                 //check for max outlier
                 //calculate border for outlier
                 #statBorderOutlier := #statQuartil75 + #rangeOutlier * #statDeltaQuartil;
                 //search in array for values outside the border 
                 FOR #statCounter := UDINT_TO_INT(#statNumberOfElements - 1) TO 0 BY -1 DO
                   #statRetVal := MOVE_BLK_VARIANT(SRC := #array, COUNT := 1, SRC_INDEX := #statCounter, DEST_INDEX := 0, DEST => #tempValueInt);
                   IF #statRetVal <> 0
                   THEN
                     #status := INT_TO_WORD(#statRetVal);
                     #statusID := #ID_INTERNAL;
                     #statError := true;
                     GOTO EndOfBlock;
                   END_IF;
                   IF #tempValueInt > #statBorderOutlier
                   THEN
                     //detected a value as outlier, check next value
                     ;
                   ELSE
                     //all outlier detected. Calulate new Max Value in range and calulate outliers in %
                     #statOutlierMax := INT_TO_REAL((100 * (UDINT_TO_INT(#statNumberOfElements) - #statCounter - 1))) / UDINT_TO_REAL(#statNumberOfElements);
                     #statMaxNew := #tempValueInt;
                     EXIT;
                   END_IF;
                 END_FOR;
               END_IF;

               //done
               #statDone := TRUE;
             END_IF;
           END_REGION ;

         ELSIF TypeOfElements(#array) = UInt
         THEN

           REGION Type is UINT
             //Type is UInt 
             //Sort array
             #instLGF_ShellSortUInt(error => #statError,
                                    statusID => #tempStatusID,
                                    status => #tempStatus,
                                    variantArray := #array);

             IF #statError = true
             THEN
               IF #tempStatusID > 1
               THEN
                 #statusID := #ID_INTERNAL;
               ELSE
                 #statusID := #ID_SORT;
                 #status := #tempStatus;
               END_IF;
               GOTO EndOfBlock;
             END_IF;

             //Identify max and min value
             #statRetVal := MOVE_BLK_VARIANT(SRC := #array, COUNT := 1, SRC_INDEX := 0, DEST_INDEX := 0, DEST => #tempMinUint);
             IF #statRetVal <> 0
             THEN
               #status := INT_TO_WORD(#statRetVal);
               #statusID := #ID_INTERNAL;
               #statError := true;
               GOTO EndOfBlock;
             END_IF;
             #statRetVal := MOVE_BLK_VARIANT(SRC := #array, COUNT := 1, SRC_INDEX := UDINT_TO_INT(#statNumberOfElements - 1), DEST_INDEX := 0, DEST => #tempMaxUint);
             IF #statRetVal <> 0
             THEN
               #status := INT_TO_WORD(#statRetVal);
               #statusID := #ID_INTERNAL;
               #statError := true;
               GOTO EndOfBlock;
             END_IF;
             #statMax := #tempMaxUint;
             #statMin := #tempMinUint;

             //calculate median (Q50)
             IF #statEven = true
             THEN
               // if n is even -> calculate MEDIAN = (x(n/2)+x(n/2+1))/2
               #statRetVal := MOVE_BLK_VARIANT(SRC := #array, COUNT := 1, SRC_INDEX := UDINT_TO_INT(#statNumberOfElements / 2), DEST_INDEX := 0, DEST => #tempValueUint);
               IF #statRetVal <> 0
               THEN
                 #status := INT_TO_WORD(#statRetVal);
                 #statusID := #ID_INTERNAL;
                 #statError := true;
                 GOTO EndOfBlock;
               END_IF;
               #statRetVal := MOVE_BLK_VARIANT(SRC := #array, COUNT := 1, SRC_INDEX := UDINT_TO_INT(#statNumberOfElements / 2) - 1, DEST_INDEX := 0, DEST => #tempValueUint1);
               IF #statRetVal <> 0
               THEN
                 #status := INT_TO_WORD(#statRetVal);
                 #statusID := #ID_INTERNAL;
                 #statError := true;
                 GOTO EndOfBlock;
               END_IF;
               #statMedian := (#tempValueUint + #tempValueUint1) / 2;
             ELSE
               // if n is odd -> MEDIAN = x(n+1/2)
               #statRetVal := MOVE_BLK_VARIANT(SRC := #array, COUNT := 1, SRC_INDEX := UDINT_TO_INT(#statNumberOfElements / 2), DEST_INDEX := 0, DEST => #tempValueUint);
               IF #statRetVal <> 0
               THEN
                 #status := INT_TO_WORD(#statRetVal);
                 #statusID := #ID_INTERNAL;
                 #statError := true;
                 GOTO EndOfBlock;
               END_IF;
               #statMedian := #tempValueUint;
             END_IF;

             //calculate 1.quartil (Q25)
             // q1 = x(k) with  k=(n+3)/4 
             #statK := (((UDINT_TO_REAL(#statNumberOfElements + 3)) / 4.0)) - 1;
             #statRetVal := MOVE_BLK_VARIANT(SRC := #array, COUNT := 1, SRC_INDEX := TRUNC(#statK), DEST_INDEX := 0, DEST => #tempValueUint);
             IF #statRetVal <> 0
             THEN
               #status := INT_TO_WORD(#statRetVal);
               #statError := true;
               GOTO EndOfBlock;
             END_IF;
             #statRetVal := MOVE_BLK_VARIANT(SRC := #array, COUNT := 1, SRC_INDEX := TRUNC(#statK) + 1, DEST_INDEX := 0, DEST => #tempValueUint1);
             IF #statRetVal <> 0
             THEN
               #status := INT_TO_WORD(#statRetVal);
               #statusID := #ID_INTERNAL;
               #statError := true;
               GOTO EndOfBlock;
             END_IF;

             #statQuartil25 := #tempValueUint + FRAC_REAL(#statK) * (#tempValueUint1 - #tempValueUint);
             //calculate 3.quartil (Q75)
             //q3 = x(n+1-k) with k=(3n+1)/4
             #statK := ((3 * UDINT_TO_REAL(#statNumberOfElements) + 1) / 4) - 1;
             #statRetVal := MOVE_BLK_VARIANT(SRC := #array, COUNT := 1, SRC_INDEX := TRUNC(#statK), DEST_INDEX := 0, DEST => #tempValueUint);
             IF #statRetVal <> 0
             THEN
               #status := INT_TO_WORD(#statRetVal);
               #statusID := #ID_INTERNAL;
               #statError := true;
               GOTO EndOfBlock;
             END_IF;
             #statRetVal := MOVE_BLK_VARIANT(SRC := #array, COUNT := 1, SRC_INDEX := TRUNC(#statK) + 1, DEST_INDEX := 0, DEST => #tempValueUint1);
             IF #statRetVal <> 0
             THEN
               #status := INT_TO_WORD(#statRetVal);
               #statusID := #ID_INTERNAL;
               #statError := true;
               GOTO EndOfBlock;
             END_IF;

             #statQuartil75 := #tempValueUint + FRAC_REAL(#statK) * (#tempValueUint1 - #tempValueUint);

             //only if RANGE_OUTLIER <> 0
             IF #rangeOutlier <> 0
             THEN

               //calculate Delta Q75-Q25
               #statDeltaQuartil := #statQuartil75 - #statQuartil25;

               //calculate border for outlier
               #statBorderOutlier := #statQuartil25 - #rangeOutlier * #statDeltaQuartil;
               //search in array for values outside the border
               FOR #statCounter := 0 TO UDINT_TO_INT(#statNumberOfElements - 1) DO
                 #statRetVal := MOVE_BLK_VARIANT(SRC := #array, COUNT := 1, SRC_INDEX := #statCounter, DEST_INDEX := 0, DEST => #tempValueUint);
                 IF #statRetVal <> 0
                 THEN
                   #status := INT_TO_WORD(#statRetVal);
                   #statusID := #ID_INTERNAL;
                   #statError := true;
                   GOTO EndOfBlock;
                 END_IF;
                 IF #tempValueUint < #statBorderOutlier
                 THEN
                   //detected a value as outlier, check next value
                   ;
                 ELSE
                   //all outlier detected. Calulate new Min Value in range and calulate outliers in %
                   #statOutlierMin := INT_TO_REAL((100 * #statCounter)) / UDINT_TO_REAL(#statNumberOfElements);
                   #statMinNew := #tempValueUint;
                   EXIT;
                 END_IF;

               END_FOR;

               //check for max outlier
               #statBorderOutlier := #statQuartil75 + #rangeOutlier * #statDeltaQuartil;

               FOR #statCounter := UDINT_TO_INT(#statNumberOfElements - 1) TO 0 BY -1 DO
                 #statRetVal := MOVE_BLK_VARIANT(SRC := #array, COUNT := 1, SRC_INDEX := #statCounter, DEST_INDEX := 0, DEST => #tempValueUint);
                 IF #statRetVal <> 0
                 THEN
                   #status := INT_TO_WORD(#statRetVal);
                   #statusID := #ID_INTERNAL;
                   #statError := true;
                   GOTO EndOfBlock;
                 END_IF;
                 IF #tempValueUint > #statBorderOutlier
                 THEN
                   //detected a value as outlier, check next value
                   ;
                 ELSE
                   //all outlier detected. Calulate new Max Value in range and calulate outliers in %
                   #statOutlierMax := INT_TO_REAL((100 * (UDINT_TO_INT(#statNumberOfElements) - #statCounter - 1))) / UDINT_TO_REAL(#statNumberOfElements);
                   #statMaxNew := #tempValueUint;
                   EXIT;
                 END_IF;
               END_FOR;
             END_IF;
             //done
             #statDone := TRUE;

           END_REGION ;

         ELSIF TypeOfElements(#array) = Real
         THEN

           REGION Type of Array is REAL

             //Type is Real
             //Sort array
             #instLGF_ShellSortReal(error => #statError,
                                    statusID => #tempStatusID,
                                    status => #tempStatus,
                                    variantArray := #array);

             IF #statError = true
             THEN
               IF #tempStatusID > 1
               THEN
                 #statusID := #ID_INTERNAL;
               ELSE
                 #statusID := #ID_SORT;
                 #status := #tempStatus;
               END_IF;
               GOTO EndOfBlock;
             END_IF;

             //Identify max and min value
             #statRetVal := MOVE_BLK_VARIANT(SRC := #array, COUNT := 1, SRC_INDEX := 0, DEST_INDEX := 0, DEST => #statMin);
             IF #statRetVal <> 0
             THEN
               #status := INT_TO_WORD(#statRetVal);
               #statusID := #ID_INTERNAL;
               #statError := true;
               GOTO EndOfBlock;
             END_IF;
             #statRetVal := MOVE_BLK_VARIANT(SRC := #array, COUNT := 1, SRC_INDEX := UDINT_TO_INT(#statNumberOfElements - 1), DEST_INDEX := 0, DEST => #statMax);
             IF #statRetVal <> 0
             THEN
               #status := INT_TO_WORD(#statRetVal);
               #statusID := #ID_INTERNAL;
               #statError := true;
               GOTO EndOfBlock;
             END_IF;

             //calculate median (Q50)
             IF #statEven = true
             THEN
               // if n is even -> calculate MEDIAN = (x(n/2)+x(n/2+1))/2
               #statRetVal := MOVE_BLK_VARIANT(SRC := #array, COUNT := 1, SRC_INDEX := UDINT_TO_INT(#statNumberOfElements / 2), DEST_INDEX := 0, DEST => #tempValueReal);
               IF #statRetVal <> 0
               THEN
                 #status := INT_TO_WORD(#statRetVal);
                 #statusID := #ID_INTERNAL;
                 #statError := true;
                 GOTO EndOfBlock;
               END_IF;
               #statRetVal := MOVE_BLK_VARIANT(SRC := #array, COUNT := 1, SRC_INDEX := UDINT_TO_INT(#statNumberOfElements / 2) - 1, DEST_INDEX := 0, DEST => #tempValueReal1);
               IF #statRetVal <> 0
               THEN
                 #status := INT_TO_WORD(#statRetVal);
                 #statusID := #ID_INTERNAL;
                 #statError := true;
                 GOTO EndOfBlock;
               END_IF;
               #statMedian := (#tempValueReal + #tempValueReal1) / 2;
             ELSE
               // if n is odd -> MEDIAN = x(n+1/2)
               #statRetVal := MOVE_BLK_VARIANT(SRC := #array, COUNT := 1, SRC_INDEX := UDINT_TO_INT(#statNumberOfElements / 2), DEST_INDEX := 0, DEST => #tempValueReal);
               IF #statRetVal <> 0
               THEN
                 #status := INT_TO_WORD(#statRetVal);
                 #statusID := #ID_INTERNAL;
                 #statError := true;
                 GOTO EndOfBlock;
               END_IF;
               #statMedian := #tempValueReal;
             END_IF;

             //calculate 1.quartil (Q25)
             // q1 = x(k) with  k=(n+3)/4 
             #statK := (((UDINT_TO_REAL(#statNumberOfElements + 3)) / 4.0)) - 1;
             #statRetVal := MOVE_BLK_VARIANT(SRC := #array, COUNT := 1, SRC_INDEX := TRUNC(#statK), DEST_INDEX := 0, DEST => #tempValueReal);
             IF #statRetVal <> 0
             THEN
               #status := INT_TO_WORD(#statRetVal);
               #statusID := #ID_INTERNAL;
               #statError := true;
               GOTO EndOfBlock;
             END_IF;
             #statRetVal := MOVE_BLK_VARIANT(SRC := #array, COUNT := 1, SRC_INDEX := TRUNC(#statK) + 1, DEST_INDEX := 0, DEST => #tempValueReal1);
             IF #statRetVal <> 0
             THEN
               #status := INT_TO_WORD(#statRetVal);
               #statusID := #ID_INTERNAL;
               #statError := true;
               GOTO EndOfBlock;
             END_IF;
             #statQuartil25 := #tempValueReal + FRAC_REAL(#statK) * (#tempValueReal1 - #tempValueReal);

             //calculate 3.quartil (Q75)
             //q3 = x(n+1-k) with k=(3n+1)/4
             #statK := ((3 * UDINT_TO_REAL(#statNumberOfElements) + 1) / 4) - 1;
             #statRetVal := MOVE_BLK_VARIANT(SRC := #array, COUNT := 1, SRC_INDEX := TRUNC(#statK), DEST_INDEX := 0, DEST => #tempValueReal);
             IF #statRetVal <> 0
             THEN
               #status := INT_TO_WORD(#statRetVal);
               #statusID := #ID_INTERNAL;
               #statError := true;
               GOTO EndOfBlock;
             END_IF;
             #statRetVal := MOVE_BLK_VARIANT(SRC := #array, COUNT := 1, SRC_INDEX := TRUNC(#statK) + 1, DEST_INDEX := 0, DEST => #tempValueReal1);
             IF #statRetVal <> 0
             THEN
               #status := INT_TO_WORD(#statRetVal);
               #statusID := #ID_INTERNAL;
               #statError := true;
               GOTO EndOfBlock;
             END_IF;
             #statQuartil75 := #tempValueReal + FRAC_REAL(#statK) * (#tempValueReal1 - #tempValueReal);

             //only if RANGE_OUTLIER <> 0
             IF #rangeOutlier <> 0
             THEN

               //calculate Delta Q75-Q25
               #statDeltaQuartil := #statQuartil75 - #statQuartil25;

               //calculate border for outlier
               #statBorderOutlier := #statQuartil25 - #rangeOutlier * #statDeltaQuartil;
               FOR #statCounter := 0 TO UDINT_TO_INT(#statNumberOfElements - 1) DO
                 #statRetVal := MOVE_BLK_VARIANT(SRC := #array, COUNT := 1, SRC_INDEX := #statCounter, DEST_INDEX := 0, DEST => #tempValueReal);
                 IF #statRetVal <> 0
                 THEN
                   #status := INT_TO_WORD(#statRetVal);
                   #statusID := #ID_INTERNAL;
                   #statError := true;
                   GOTO EndOfBlock;
                 END_IF;
                 IF #tempValueReal < #statBorderOutlier
                 THEN
                   //detected a value as outlier, check next value
                   ;
                 ELSE
                   //all outlier detected. Calulate new Min Value in range and calulate outliers in %
                   #statOutlierMin := INT_TO_REAL((100 * #statCounter)) / UDINT_TO_REAL(#statNumberOfElements);
                   #statMinNew := #tempValueReal;
                   EXIT;
                 END_IF;

               END_FOR;

               //check for max outlier
               //calculate border for outlier
               #statBorderOutlier := #statQuartil75 + #rangeOutlier * #statDeltaQuartil;
               FOR #statCounter := UDINT_TO_INT(#statNumberOfElements - 1) TO 0 BY -1 DO
                 #statRetVal := MOVE_BLK_VARIANT(SRC := #array, COUNT := 1, SRC_INDEX := #statCounter, DEST_INDEX := 0, DEST => #tempValueReal);
                 IF #statRetVal <> 0
                 THEN
                   #status := INT_TO_WORD(#statRetVal);
                   #statusID := #ID_INTERNAL;
                   #statError := true;
                   GOTO EndOfBlock;
                 END_IF;
                 IF #tempValueReal > #statBorderOutlier
                 THEN
                   //detected a value as outlier, check next value
                   ;
                 ELSE
                   //all outlier detected. Calulate new Max Value in range and calulate outliers in %
                   #statOutlierMax := INT_TO_REAL((100 * (UDINT_TO_INT(#statNumberOfElements) - #statCounter - 1))) / UDINT_TO_REAL(#statNumberOfElements);
                   #statMaxNew := #tempValueReal;
                   EXIT;
                 END_IF;
               END_FOR;
             END_IF;
             //done
             #statDone := TRUE;

           END_REGION ;

         ELSE
           #statError := true;
           #status := #STATUS_WRONG_DATATYPE;
         END_IF;
         //calculate Skewness
         //S= ((Q25 + Q75)-2*Q50) / (Q75 - Q25)
         #skewness := (#statQuartil75 + #statQuartil25 - 2.0 * #statMedian) / (#statQuartil75 - #statQuartil25);

         //write output values
         IF #rangeOutlier <> 0
         THEN
           #min := #statMinNew;
           #max := #statMaxNew;
         ELSE
           #min := #statMin;
           #max := #statMax;
         END_IF;

         #q25 := #statQuartil25;
         #median := #statMedian;
         #q75 := #statQuartil75;
         #outlierMin := #statOutlierMin;
         #outlierMax := #statOutlierMax;
         GOTO EndOfBlock;

       END_IF;
     ELSE
       #statError := true;
       #status := #STATUS_NO_ARRAY;
     END_IF;


   END_REGION

   REGION Write Outputs
     //Error occured in request


   EndOfBlock:
     IF #statError
     THEN
       #statDone := FALSE;
       #statBusy := FALSE;
       //Request finished
     ELSIF #statDone
     THEN
       #statBusy := FALSE;
       #statError := FALSE;
       #status := #STATUS_EXECUTION_FINISHED;

       //Request in execution
     ELSE
       #status := #STATUS_SUBSEQUENT_CALL;
     END_IF;


     //Write static values (done,busy,error) to outputs
     #done := #statDone;
     #busy := #statBusy;
     #error := #statError;
     //----------------------------------------------------------------------------------------------

   END_REGION ;
END_FUNCTION_BLOCK

FUNCTION_BLOCK "LGF_Histogram"   // FB10011, SCL
{ S7_Optimized_Access := 'TRUE' }
VERSION : 0.1
   VAR_INPUT
      execute : Bool;   // Rising edge starts action once
      NumberOfClasses : UInt;   // Number of desired classes.
   END_VAR
   VAR_OUTPUT
      busy : Bool;   // TRUE: FB is not finished and new output values can be expected
      done : Bool;   // TRUE: Commanded action has been completed successfully
      error : Bool;   // Rising edge informs that an error occurred during the execution of
      status : Word := 16#7000;   // Current status of FB
      statusID : UInt := 1;   // Current statusID of FB
      histValues : Array[0..1, 0..14] of Real;   // Outputs the calculated values in a two-dimensional array
      axis : Array[0..3] of Real;   // Specifies the axis values
      classWidth : Real;   // Returns the calculated class width.
   END_VAR
   VAR_IN_OUT
      "array" : Variant;
   END_VAR
   VAR
      statBusy : Bool;   // Static value for output busy
      statDone : Bool;   // Static value for output done
      statError : Bool;   // Static value for output error
      statExecuteOld : Bool;   // Old value of execute for edge detection
      instLGF_ShellSortInt : "LGF_ShellSortInt";   // Instance of LG_ShellSortInt
      instLGF_ShellSortReal : "LGF_ShellSortReal";   // Instance of LG_ShellSortReal
      instLGF_ShellSortUInt : "LGF_ShellSortUInt";   // Instance of LG_ShellSortUInt
      statMin : Real;   // Static value for min
      statMax : Real;   // Static value for max
      statNumberOfElements : UDInt;   // Static value for number of elements
      statType : Int;   // Static value for type
      statAverage : Real;   // Static value for average
      statDeviation : Real;   // Static value for deviation
      statCounter : Int;   // Static value for counter
      statWidth : Real;   // Static value for width
      statFrequencyValues : Int;   // Static value for frequency values
      statI : Int;   // Static value for I
      statIold : Int := 0;   // Static value for I old
      statBound : Real;   // Static value for bound
      statMaxFrequency : Int;   // Static value for max frequency
      statHistFrequencyAbs : Array[0..14] of Int;   // Static array for history frequency absolute
      statHistFrequencyRel : Array[0..14] of Real;   // Static array for history frequency relative
      statHistMiddleOfClass : Array[0..14] of Real;   // Static array for history middle of class
   END_VAR
   VAR_TEMP
      tempError : Bool;   // Temporary error
      tempStatusID : UInt;   // Temporary status ID
      tempStatus : Word;   // Temporary status
      tempRetVal : Int;   // Temporary RetVal
      tempValueInt : Int;   // Temporary value for calculation
      tempValueUint : UInt;   // Temporary value for calculation
      tempValueReal : Real;   // Temporary value for calculation
      tempMinInt : Int;   // Temporary value for min INT
      tempMaxInt : Int;   // Temporary value for max INT
      tempMinUint : UInt;   // Temporary value for min UINT
      tempMaxUint : UInt;   // Temporary value for max UINT
   END_VAR
   VAR CONSTANT
      STATUS_EXECUTION_FINISHED : Word := 16#0000;   // Status: Execution finished without errors
      STATUS_NO_CALL : Word := 16#7000;   // Status: No call of FB
      STATUS_FIRST_CALL : Word := 16#7001;   // Status: First call of FB after enabling
      STATUS_SUBSEQUENT_CALL : Word := 16#7002;   // Status: Subsequent call of FB
      STATUS_WRONG_DATATYPE : Word := 16#9100;   // Status: Wrong data type
      STATUS_WRONG_NO_CLASSES : Word := 16#9101;   // Status: Wrong number of classes
      STATUS_NO_ARRAY : Word := 16#9102;   // Status: No array
      TYPE_INT : Int := 0;   // TYPE: INT
      TYPE_UINT : Int := 1;   // TYPE: UINT
      TYPE_REAL : Int := 2;   // TYPE: REAL
      ID_INTERNAL : UInt := 1;   // Status ID: Internal error
      ID_MOVE_BLK : UInt := 2;   // Status ID: Function MOVE_BLK
      ID_SORT : UInt := 3;   // Status ID: Error sorting
   END_VAR
BEGIN
   //=============================================================================
   // SIEMENS AG
   // (c)Copyright 2017
   //-----------------------------------------------------------------------------
   // Library:       LGF (Library General Functions)
   // Tested with:   CPU1212C DC/DC/DC FW:V4.2
   // Engineering:   TIA Portal V15.1 
   // Restrictions:  -
   // Requirements:  PLC (S7-1200 / S7-1500)
   // Functionality: calculate from measurement list all values for creating
   //                a histogramm with WinCC
   //-----------------------------------------------------------------------------
   // Change log table:
   // Version  Date        In charge / Changes applied
   // 01.00.00 23.11.2018  Siemens Industry Online Support
   //                      First released version
   //=============================================================================

   //Check if FB is triggered
   //Too many classes on input. MAX = 15 Classes

   //FB is active
   IF #execute
     AND NOT #statExecuteOld
     AND NOT #statBusy
   THEN
     //Functionality is busy
     #statBusy := TRUE;

     //Reset other outputs
     #statError := FALSE;
     #status := #STATUS_FIRST_CALL;

     //Reset statics
     FILL_BLK(IN := 0,
              COUNT := 15,
              OUT => #statHistFrequencyAbs[0]);
     FILL_BLK(IN := 0,
              COUNT := 15,
              OUT => #statHistFrequencyRel[0]);
     FILL_BLK(IN := 0,
              COUNT := 15,
              OUT => #statHistMiddleOfClass[0]);
     #statI := 0;
     #statFrequencyValues := 0;
     #statIold := 0;

     #statExecuteOld := #execute;
     #statMaxFrequency := 0;

     GOTO EndOfBlock;
     //FB is currently inactive
   ELSIF NOT #execute
     AND NOT #statBusy
   THEN
     //Error outputs are reset with falling edge of enable input
     #statError := FALSE;

     //Done and busy are reset with falling edge of enable input
     #statDone := FALSE;
     #statBusy := FALSE;

     //Write outputs
     #status := #STATUS_NO_CALL;
     #statExecuteOld := #execute;

     GOTO EndOfBlock;
     //FB is currently executed and not finished
   ELSIF #statBusy
   THEN
     #statExecuteOld := #execute;

     //FB finished job
   ELSE
     #statExecuteOld := #execute;
     //Wait for start of functionality 
   END_IF;

   IF #statBusy = true
     AND #statError = false
   THEN

     REGION check Datatype of Array, sort and count the elements

       //count array elements
       #statNumberOfElements := CountOfElements(#array);

       //check number of classes
       IF (#NumberOfClasses > 15)
         OR (#NumberOfClasses < 1)
       THEN
         #statError := true;
         #status := #STATUS_WRONG_NO_CLASSES;
         #statusID := #ID_INTERNAL;
         GOTO EndOfBlock;
       END_IF;

       IF IS_ARRAY(#array)
       THEN
         //check which datatype is used
         IF TypeOfElements(#array) = Int
         THEN
           //Type is Int
           REGION Type of Array is INT
             //Sort array
             #instLGF_ShellSortInt(error => #statError,
                                   statusID => #tempStatusID,
                                   status => #tempStatus,
                                   variantArray := #array);
             IF #statError = true
             THEN
               IF #tempStatusID > 1
               THEN
                 #statusID := #ID_INTERNAL;
               ELSE
                 #statusID := #ID_SORT;
               END_IF;
               #status := #tempStatus;
               GOTO EndOfBlock;
             ELSE
               //Identify max and min value
               #tempRetVal := MOVE_BLK_VARIANT(SRC := #array, COUNT := 1, SRC_INDEX := 0, DEST_INDEX := 0, DEST => #tempMinInt);
               IF #tempRetVal <> 0
               THEN
                 #status := INT_TO_WORD(#tempRetVal);
                 #statusID := #ID_MOVE_BLK;
                 #statError := true;
                 GOTO EndOfBlock;
               END_IF;
               #tempRetVal := MOVE_BLK_VARIANT(SRC := #array, COUNT := 1, SRC_INDEX := UDINT_TO_INT(#statNumberOfElements - 1), DEST_INDEX := 0, DEST => #tempMaxInt);
               IF #tempRetVal <> 0
               THEN
                 #status := INT_TO_WORD(#tempRetVal);
                 #statusID := #ID_MOVE_BLK;
                 #statError := true;
                 GOTO EndOfBlock;
               END_IF;

               #statMin := INT_TO_REAL(#tempMinInt);
               #statMax := INT_TO_REAL(#tempMaxInt);

               //calculate classwidth
               #statWidth := (#statMax - #statMin) / #NumberOfClasses;
               #statBound := (#statMin + #statWidth);

               //search for all values
               FOR #statCounter := 0 TO UINT_TO_INT(#NumberOfClasses) - 1 DO

                 //Count Values for Class 
                 #tempRetVal := MOVE_BLK_VARIANT(SRC := #array, COUNT := 1, SRC_INDEX := 0, DEST_INDEX := 0, DEST => #tempValueInt);
                 IF #tempRetVal <> 0
                 THEN
                   #status := INT_TO_WORD(#tempRetVal);
                   #statusID := #ID_MOVE_BLK;
                   #statError := true;
                   GOTO EndOfBlock;
                 END_IF;
                 WHILE (#tempValueInt < #statBound)
                   AND #statI < #statNumberOfElements - 1 DO

                   IF #statI = #statNumberOfElements
                   THEN
                     EXIT;
                   END_IF;
                   #statI := #statI + 1;
                   #tempRetVal := MOVE_BLK_VARIANT(SRC := #array, COUNT := 1, SRC_INDEX := #statI, DEST_INDEX := 0, DEST => #tempValueInt);
                   IF #tempRetVal <> 0
                   THEN
                     #status := INT_TO_WORD(#tempRetVal);
                     #statusID := #ID_MOVE_BLK;
                     #statError := true;
                     GOTO EndOfBlock;
                   END_IF;
                 END_WHILE;

                 //the last value is not counted, because of rounding errors
                 IF #statI = #statNumberOfElements - 1
                 THEN
                   #statI := #statI + 1;
                 END_IF;

                 #statFrequencyValues := #statI - #statIold;
                 #statHistFrequencyAbs[#statCounter] := #statFrequencyValues;

                 #statHistFrequencyRel[#statCounter] := INT_TO_REAL(#statFrequencyValues) / UDINT_TO_REAL(#statNumberOfElements) * 100;

                 //Max values in one class for y-axis 
                 IF #statMaxFrequency < #statFrequencyValues
                 THEN
                   #statMaxFrequency := #statFrequencyValues;
                 END_IF;

                 #statBound := #statBound + #statWidth;
                 #statIold := #statI;
               END_FOR;
             END_IF;
           END_REGION

         ELSIF TypeOfElements(#array) = UInt
         THEN
           //Type is UInt 
           REGION Type of Array is UINT
             //Sort array
             #instLGF_ShellSortUInt(error => #statError,
                                    statusID => #tempStatusID,
                                    status => #tempStatus,
                                    variantArray := #array);
             IF #statError = true
             THEN
               IF #tempStatusID > 1
               THEN
                 #statusID := #ID_INTERNAL;
               ELSE
                 #statusID := #ID_SORT;
               END_IF;
               #status := #tempStatus;
               GOTO EndOfBlock;
             ELSE
               //Identify max and min value
               #tempRetVal := MOVE_BLK_VARIANT(SRC := #array, COUNT := 1, SRC_INDEX := 0, DEST_INDEX := 0, DEST => #tempMinUint);
               IF #tempRetVal <> 0
               THEN
                 #status := INT_TO_WORD(#tempRetVal);
                 #statusID := #ID_MOVE_BLK;
                 #statError := true;
                 GOTO EndOfBlock;
               END_IF;
               #tempRetVal := MOVE_BLK_VARIANT(SRC := #array, COUNT := 1, SRC_INDEX := UDINT_TO_INT(#statNumberOfElements - 1), DEST_INDEX := 0, DEST => #tempMaxUint);
               IF #tempRetVal <> 0
               THEN
                 #status := INT_TO_WORD(#tempRetVal);
                 #statusID := #ID_MOVE_BLK;
                 #statError := true;
                 GOTO EndOfBlock;
               END_IF;

               #statMin := UINT_TO_REAL(#tempMinUint);
               #statMax := UINT_TO_REAL(#tempMaxUint);

               //calculate classwidth
               #statWidth := (#statMax - #statMin) / #NumberOfClasses;
               #statBound := (#statMin + #statWidth);

               //search for all values
               FOR #statCounter := 0 TO UINT_TO_INT(#NumberOfClasses) - 1 DO

                 //Count Values for Class 
                 #tempRetVal := MOVE_BLK_VARIANT(SRC := #array, COUNT := 1, SRC_INDEX := 0, DEST_INDEX := 0, DEST => #tempValueUint);
                 IF #tempRetVal <> 0
                 THEN
                   #status := INT_TO_WORD(#tempRetVal);
                   #statusID := #ID_MOVE_BLK;
                   #statError := true;
                   GOTO EndOfBlock;

                 END_IF;
                 WHILE (#tempValueUint < #statBound)
                   AND #statI < #statNumberOfElements - 1 DO

                   IF #statI = #statNumberOfElements
                   THEN
                     EXIT;
                   END_IF;
                   #statI := #statI + 1;
                   #tempRetVal := MOVE_BLK_VARIANT(SRC := #array, COUNT := 1, SRC_INDEX := #statI, DEST_INDEX := 0, DEST => #tempValueUint);
                   IF #tempRetVal <> 0
                   THEN
                     #status := INT_TO_WORD(#tempRetVal);
                     #statusID := #ID_MOVE_BLK;
                     #statError := true;
                     GOTO EndOfBlock;
                   END_IF;
                 END_WHILE;

                 //the last value is not counted, because of rounding errors
                 IF #statI = #statNumberOfElements - 1
                 THEN
                   #statI := #statI + 1;
                 END_IF;

                 #statFrequencyValues := #statI - #statIold;
                 #statHistFrequencyAbs[#statCounter] := #statFrequencyValues;

                 #statHistFrequencyRel[#statCounter] := INT_TO_REAL(#statFrequencyValues) / UDINT_TO_REAL(#statNumberOfElements) * 100;

                 //Max values in one class for y-axis 
                 IF #statMaxFrequency < #statFrequencyValues
                 THEN
                   #statMaxFrequency := #statFrequencyValues;
                 END_IF;

                 #statBound := #statBound + #statWidth;
                 #statIold := #statI;
               END_FOR;

             END_IF;
           END_REGION

         ELSIF TypeOfElements(#array) = Real
         THEN
           //Type is Real
           REGION Type of Array is REAL
             //Sort array
             #instLGF_ShellSortReal(error => #statError,
                                    statusID => #tempStatusID,
                                    status => #tempStatus,
                                    variantArray := #array);
             IF #statError = true
             THEN
               IF #tempStatusID > 1
               THEN
                 #statusID := #ID_INTERNAL;
               ELSE
                 #statusID := #ID_SORT;
               END_IF;
               #status := #tempStatus;
               GOTO EndOfBlock;
             ELSE
               //Identify max and min value
               #tempRetVal := MOVE_BLK_VARIANT(SRC := #array, COUNT := 1, SRC_INDEX := 0, DEST_INDEX := 0, DEST => #statMin);
               IF #tempRetVal <> 0
               THEN
                 #status := INT_TO_WORD(#tempRetVal);
                 #statusID := #ID_MOVE_BLK;
                 #statError := true;
                 GOTO EndOfBlock;
               END_IF;
               #tempRetVal := MOVE_BLK_VARIANT(SRC := #array, COUNT := 1, SRC_INDEX := UDINT_TO_INT(#statNumberOfElements - 1), DEST_INDEX := 0, DEST => #statMax);
               IF #tempRetVal <> 0
               THEN
                 #status := INT_TO_WORD(#tempRetVal);
                 #statusID := #ID_MOVE_BLK;
                 #statError := true;
                 GOTO EndOfBlock;
               END_IF;
               //calculate classwidth
               #statWidth := (#statMax - #statMin) / #NumberOfClasses;
               #statBound := (#statMin + #statWidth);

               //search for all values
               FOR #statCounter := 0 TO UINT_TO_INT(#NumberOfClasses) - 1 DO

                 //Count Values for Class 
                 #tempRetVal := MOVE_BLK_VARIANT(SRC := #array, COUNT := 1, SRC_INDEX := 0, DEST_INDEX := 0, DEST => #tempValueReal);
                 IF #tempRetVal <> 0
                 THEN
                   #status := INT_TO_WORD(#tempRetVal);
                   #statusID := #ID_MOVE_BLK;
                   #statError := true;
                   GOTO EndOfBlock;
                 END_IF;
                 WHILE (#tempValueReal < #statBound)
                   AND #statI < #statNumberOfElements - 1 DO

                   IF #statI = #statNumberOfElements
                   THEN
                     EXIT;
                   END_IF;
                   #statI := #statI + 1;
                   #tempRetVal := MOVE_BLK_VARIANT(SRC := #array, COUNT := 1, SRC_INDEX := #statI, DEST_INDEX := 0, DEST => #tempValueReal);
                   IF #tempRetVal <> 0
                   THEN
                     #status := INT_TO_WORD(#tempRetVal);
                     #statusID := #ID_MOVE_BLK;
                     #statError := true;
                     GOTO EndOfBlock;
                   END_IF;
                 END_WHILE;

                 //the last value is not counted, because of rounding errors
                 IF #statI = #statNumberOfElements - 1
                 THEN
                   #statI := #statI + 1;
                 END_IF;

                 #statFrequencyValues := #statI - #statIold;
                 #statHistFrequencyAbs[#statCounter] := #statFrequencyValues;
                 #statHistFrequencyRel[#statCounter] := INT_TO_REAL(#statFrequencyValues) / UDINT_TO_REAL(#statNumberOfElements) * 100;

                 //Max values in one class for y-axis 
                 IF #statMaxFrequency < #statFrequencyValues
                 THEN
                   #statMaxFrequency := #statFrequencyValues;
                 END_IF;

                 #statBound := #statBound + #statWidth;
                 #statIold := #statI;
               END_FOR;
             END_IF;
             #statDone := true;
           END_REGION

         ELSE
           #statError := true;
           #status := #STATUS_WRONG_DATATYPE;
           GOTO EndOfBlock;
         END_IF;
       ELSE
         #statError := true;
         #status := #STATUS_NO_ARRAY;
         GOTO EndOfBlock;
       END_IF;

       //find the middle of each class
       FOR #statCounter := 0 TO UINT_TO_INT(#NumberOfClasses) - 1 DO
         #statHistMiddleOfClass[#statCounter] := #statMin + (DINT_TO_REAL(#statCounter) * #statWidth) + #statWidth / 2;
       END_FOR;

       //calculate Axis values
       #axis[0] := #statMin;
       #axis[1] := #statMax;
       #axis[2] := 0.0;
       #axis[3] := INT_TO_REAL(#statMaxFrequency);

       //write class width
       #classWidth := #statWidth;

       //copy values to output array
       FOR #statCounter := 0 TO 14 DO
         #histValues[0, #statCounter] := #statHistFrequencyRel[#statCounter];
         #histValues[1, #statCounter] := #statHistMiddleOfClass[#statCounter];
       END_FOR;

     END_REGION

   END_IF;

   EndOfBlock:
   //----------------------------------------------------------------------------------------------
   //Write ouputs and error handling
   //----------------------------------------------------------------------------------------------
   //Error occured in request
   IF #statError
   THEN
     #statDone := FALSE;
     #statBusy := FALSE;
     //Request finished
   ELSIF #statDone
   THEN
     #statBusy := FALSE;
     #statError := FALSE;
     #status := #STATUS_EXECUTION_FINISHED;
     #statusID := #ID_INTERNAL;
     //Request in execution
   ELSE
     #status := #STATUS_SUBSEQUENT_CALL;
   END_IF;

   //Write static values to outputs
   #done := #statDone;
   #busy := #statBusy;
   #error := #statError;
   //----------------------------------------------------------------------------------------------
END_FUNCTION_BLOCK

FUNCTION_BLOCK "LGF_SmoothByPolynomFB"   // FB10013, SCL
{ S7_Optimized_Access := 'TRUE' }
VERSION : 0.1
   VAR_INPUT
      enable : Bool;   // TRUE: Enable functionality of FB; 0: Disable
      insert : Bool;   // Positive edge inserts a new value
      value : Real;   // The value
   END_VAR
   VAR_OUTPUT
      smoothedValue : Real;   // The smoothed value
      busy : Bool;   // TRUE: FB is working and new output values can be expected
      valid : Bool;   // TRUE: Valid set of outputs available at the FB
      error : Bool;   // Rising edge informs that an error occurred during the execution of
      status : Word := 16#7000;   // Current status of FB
   END_VAR
   VAR
      statErrorUserCleared : Bool;   // Error occured that can only be solved by user; rising edge at enable input necessary
      statErrorAutoCleared : Bool;   // Error occured that can be acknowledged by FB
      statEnableOld : Bool;   // Old value of enable for edge detection
      statValues : Array[0..4] of Real;   // Static array values
      statCount : Int;   // Static value for count
      statNoValues : Bool;   // Static value for no values
      statInsertOld : Bool;   // Static value for insert
   END_VAR
   VAR CONSTANT
      STATUS_EXECUTION_FINISHED : Word := 16#0000;   // Status: Execution finished without errors
      STATUS_NO_CALL : Word := 16#7000;   // Status: No call of FB
      STATUS_FIRST_CALL : Word := 16#7001;   // Status: First call of FB after enabling
      STATUS_SUBSEQUENT_CALL : Word := 16#7002;   // Status: Subsequent call of FB
      STATUS_NOT_ENOUGH_VALUES : Word := 16#9000;   // Status: Not enough values (3 values needed)
   END_VAR
BEGIN
   //=============================================================================
   // SIEMENS AG
   // (c)Copyright 2018
   //-----------------------------------------------------------------------------
   // Library:       LGF (Library General Functions)
   // Tested with:   CPU1212C DC/DC/DC FW:V4.2
   // Engineering:   TIA Portal V15.1 
   // Restrictions:  -
   // Requirements:  PLC (S7-1200 / S7-1500)
   // Functionality: This function block calculates the smoothed values 
   //-----------------------------------------------------------------------------
   // Change log table:
   // Version  Date        In charge / Changes applied
   // 01.00.00 23.11.2018  Siemens Industry Online Support
   //                      First released version
   //=============================================================================

   //Check if FB is disabled
   IF NOT #enable
     AND #statEnableOld
   THEN

     //Error outputs are reset with falling edge of enable input
     #statErrorUserCleared := FALSE;
     #statErrorAutoCleared := FALSE;
     #error := FALSE;
     #status := #STATUS_NO_CALL;

     //Enable and busy are reset with falling edge of enable input
     #valid := FALSE;
     #busy := FALSE;

     //Set old value of enable for edge detection and end execution
     #statEnableOld := #enable;
     RETURN;

     //Check if FB is enabled
   ELSIF #enable
     AND NOT #statEnableOld
   THEN
     //reset static values
     #statCount := 0;
     #statValues[0] := 0.0;
     #statValues[1] := 0.0;
     #statValues[2] := 0.0;
     #statValues[3] := 0.0;
     #statValues[4] := 0.0;

     #smoothedValue := 0.0;
     #statNoValues := true;

     //Busy is set at rising edge of enable input
     #busy := TRUE;
     //Set status for first call
     #status := #STATUS_FIRST_CALL;
     //Set old value of enable for edge detection and end execution
     #statEnableOld := #enable;
     RETURN;

     //Check if user cleared error in FB occurred
   ELSIF #statErrorUserCleared


   THEN
     #busy := FALSE;
     //Set old value of enable for edge detection and end execution
     #statEnableOld := #enable;
     //No set of status necessary, because status already set when error occured
     RETURN;

     //Check if function block is disabled
   ELSIF NOT #enable
   THEN
     #busy := FALSE;
     #status := #STATUS_NO_CALL;
     //Set old value of enable for edge detection and end execution
     #statEnableOld := #enable;
     RETURN;

   ELSE
     //Detect edge for disabling
     #statEnableOld := #enable;
   END_IF;


   //----------------------------------------------------------------------------------------------
   //set Status "Not enough values" after reset
   IF #enable
     AND #statEnableOld
     AND #statNoValues
   THEN
     #status := #STATUS_NOT_ENOUGH_VALUES;
     #statErrorAutoCleared := true;
     #statNoValues := false;
   END_IF;

   // positive edge of insert detected 
   IF #insert
     AND NOT #statInsertOld
   THEN

     #statInsertOld := #insert;

     #statValues[0] := #statValues[1]; // -> n-2
     #statValues[1] := #statValues[2]; // -> n-1
     #statValues[2] := #statValues[3]; // -> n
     #statValues[3] := #statValues[4]; // -> n+1
     #statValues[4] := #value;         // -> n+2

     IF #statCount < 4 THEN
       #statCount += 1;
       #status := #STATUS_NOT_ENOUGH_VALUES;
       #statErrorAutoCleared := true;
     ELSE
       //calculate new smoothed value 
       //y(n)=1/35*(-3*y(n-2)+12*y(n-1)+17*y(n)+12*y(n+1)-3*y(n+2))
       //1/35 = 0.028571
       #smoothedValue := 0.028571 * (-3 * #statValues[0] + 12 * #statValues[1] + 17 * #statValues[2] + 12 * #statValues[3] - 3 * #statValues[4]);
     END_IF;
   ELSE

     #statInsertOld := #insert;
   END_IF;

   //----------------------------------------------------------------------------------------------
   //Error handling 
   //----------------------------------------------------------------------------------------------
   IF #statErrorUserCleared
   THEN
     #valid := FALSE;
     #busy := FALSE;
     #error := TRUE;

     RETURN;

   ELSIF #statErrorAutoCleared
   THEN
     #valid := FALSE;
     #busy := TRUE;
     #error := TRUE;

     RETURN;

   ELSE
     //Process normal output values
     #valid := TRUE;
     #error := FALSE;
     #status := #STATUS_SUBSEQUENT_CALL; //Set status for subsequent call
   END_IF;
   //----------------------------------------------------------------------------------------------
END_FUNCTION_BLOCK

FUNCTION_BLOCK "LGF_DifferenceQuotientFB"   // FB10014, SCL
{ S7_Optimized_Access := 'TRUE' }
VERSION : 0.1
   VAR_INPUT
      enable : Bool;   // Activates the block. As long as "enable" is "true", the block can accept values at the "value" parameter.
      insert : Bool;   // Accepts the value at input "value" and outputs a "derivatedValue" if five values have been read in.
      value : Real;   // Value that is to be included in the differentiation.
      deltaT : Real;   // Equidistant distance between two measured values. (e.g. 1s)
   END_VAR
   VAR_OUTPUT
      derivatedValue : Real;   // Differentiated value.
      busy : Bool;   // Processing of the block is active.
      valid : Bool;   // Processing was completed successfully.
      error : Bool;   // An error occurred during processing.
      status : Word;   // Outputs the status code of the processing
   END_VAR
   VAR
      statErrorUserCleared : Bool;   // Error occured that can only be solved by user; rising edge at enable input necessary
      statErrorAutoCleared : Bool;   // Error occured that can be acknowledged by FB
      statEnableOld : Bool;   // Old value of enable for edge detection
      statDone : Bool;   // Static value for done
      statValues : Array[0..4] of Real;   // Static array values
      statCount : Int;   // Static value for count
      statDerivatedValue : Real;   // Static derivated value
      statNoValues : Bool;   // Static value for no values
      statInsertOld : Bool;   // Static value for insert
   END_VAR
   VAR CONSTANT
      STATUS_EXECUTION_FINISHED : Word := 16#0000;   // Status: Execution finished without errors
      STATUS_NO_CALL : Word := 16#7000;   // Status: No call of FB
      STATUS_FIRST_CALL : Word := 16#7001;   // Status: First call of FB after enabling
      STATUS_SUBSEQUENT_CALL : Word := 16#7002;   // Status: Subsequent call of FB
      STATUS_NOT_ENOUGH_VALUES : Word := 16#9000;   // Status: Not enough values. 5 values needed
   END_VAR
BEGIN
   //=============================================================================
   // SIEMENS AG
   // (c)Copyright 2017
   //-----------------------------------------------------------------------------
   // Library:       LGF (Library General Functions)
   // Tested with:   CPU1212C DC/DC/DC FW:V4.2
   // Engineering:   TIA Portal V15.1 
   // Restrictions:  -
   // Requirements:  PLC (S7-1200 / S7-1500)
   // Functionality: This function block differentiates a signal 
   //-----------------------------------------------------------------------------
   // Change log table:
   // Version  Date        In charge / Changes applied
   // 01.00.00 23.11.2018  Siemens Industry Online Support
   //                      First released version
   //=============================================================================

   //Check if FB is triggered
   IF #enable
       AND NOT #statEnableOld
       AND NOT #statErrorUserCleared
   THEN
       //Functionality is busy
       #statErrorUserCleared := TRUE;

       //Reset other outputs
       #statErrorAutoCleared := FALSE;
       #status := #STATUS_FIRST_CALL;

       //Reset 
   ELSIF #insert
   THEN

       #statCount := 0;

       #statValues[0] := 0.0;
       #statValues[1] := 0.0;
       #statValues[2] := 0.0;
       #statValues[3] := 0.0;
       #statValues[4] := 0.0;

       #derivatedValue := 0.0;

       #statEnableOld := #enable;

       //FB is currently inactive
   ELSIF NOT #enable
       AND NOT #statErrorUserCleared
   THEN
       //Error outputs are reset with falling edge of enable input
       #statErrorAutoCleared := FALSE;

       //Done and busy are reset with falling edge of enable input
       #statDone := FALSE;
       #statErrorUserCleared := FALSE;

       //Write outputs
       #status := #STATUS_NO_CALL;

       #statEnableOld := #enable;
   END_IF;
       //FB is currently executed and not finished
   IF #statErrorUserCleared
   THEN
       #statEnableOld := #enable;

       //FB finished job
   ELSE
       #statEnableOld := #enable;
       //Wait for start of functionality 
   END_IF;
   //----------------------------------------------------------------------------------------------